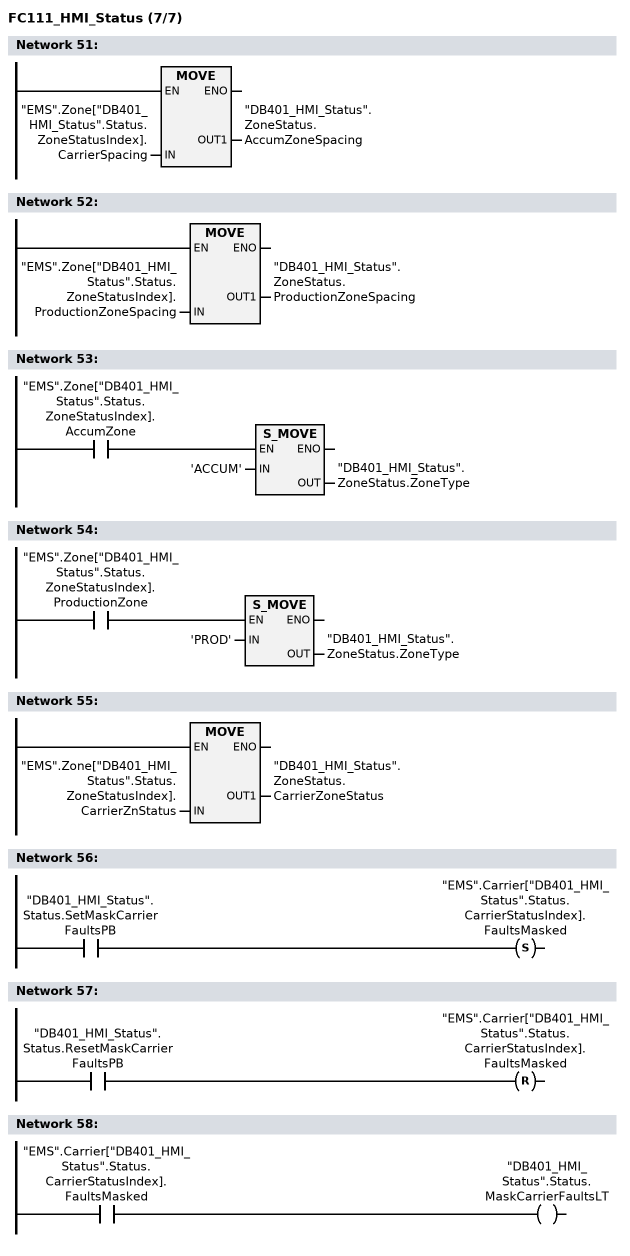
   RUNG wire#powerrail
      Move(in := "EMS".Zone["DB401_HMI_Status".Status.ZoneStatusIndex].CarrierSpacing, out1 => "DB401_HMI_Status".ZoneStatus.AccumZoneSpacing)
   END_RUNG
   // the same network as SCL:
   "DB401_HMI_Status".ZoneStatus.AccumZoneSpacing := "EMS".Zone["DB401_HMI_Status".Status.ZoneStatusIndex].CarrierSpacing;
END_REGION

REGION Network 52
   RUNG wire#powerrail
      Move(in := "EMS".Zone["DB401_HMI_Status".Status.ZoneStatusIndex].ProductionZoneSpacing, out1 => "DB401_HMI_Status".ZoneStatus.ProductionZoneSpacing)
   END_RUNG
   // the same network as SCL:
   "DB401_HMI_Status".ZoneStatus.ProductionZoneSpacing := "EMS".Zone["DB401_HMI_Status".Status.ZoneStatusIndex].ProductionZoneSpacing;
END_REGION

REGION Network 53
   RUNG wire#powerrail
      Contact( "EMS".Zone["DB401_HMI_Status".Status.ZoneStatusIndex].AccumZone )
      S_Move(in := 'ACCUM', out => "DB401_HMI_Status".ZoneStatus.ZoneType)
   END_RUNG
   // the same network as SCL:
   IF "EMS".Zone["DB401_HMI_Status".Status.ZoneStatusIndex].AccumZone THEN
       "DB401_HMI_Status".ZoneStatus.ZoneType := 'ACCUM';
   END_IF;
END_REGION

REGION Network 54
   RUNG wire#powerrail
      Contact( "EMS".Zone["DB401_HMI_Status".Status.ZoneStatusIndex].ProductionZone )
      S_Move(in := 'PROD', out => "DB401_HMI_Status".ZoneStatus.ZoneType)
   END_RUNG
   // the same network as SCL:
   IF "EMS".Zone["DB401_HMI_Status".Status.ZoneStatusIndex].ProductionZone THEN
       "DB401_HMI_Status".ZoneStatus.ZoneType := 'PROD';
   END_IF;
END_REGION

REGION Network 55
   RUNG wire#powerrail
      Move(in := "EMS".Zone["DB401_HMI_Status".Status.ZoneStatusIndex].CarrierZnStatus, out1 => "DB401_HMI_Status".ZoneStatus.CarrierZoneStatus)
   END_RUNG
   // the same network as SCL:
   "DB401_HMI_Status".ZoneStatus.CarrierZoneStatus := "EMS".Zone["DB401_HMI_Status".Status.ZoneStatusIndex].CarrierZnStatus;
END_REGION

REGION Network 56
   RUNG wire#powerrail
      Contact( "DB401_HMI_Status".Status.SetMaskCarrierFaultsPB )
      S_Coil( "EMS".Carrier["DB401_HMI_Status".Status.CarrierStatusIndex].FaultsMasked )
   END_RUNG
   // the same network as SCL:
   IF "DB401_HMI_Status".Status.SetMaskCarrierFaultsPB THEN
       "EMS".Carrier["DB401_HMI_Status".Status.CarrierStatusIndex].FaultsMasked := TRUE;
   END_IF;
END_REGION

REGION Network 57
   RUNG wire#powerrail
      Contact( "DB401_HMI_Status".Status.ResetMaskCarrierFaultsPB )
      R_Coil( "EMS".Carrier["DB401_HMI_Status".Status.CarrierStatusIndex].FaultsMasked )
   END_RUNG
   // the same network as SCL:
   IF "DB401_HMI_Status".Status.ResetMaskCarrierFaultsPB THEN
       "EMS".Carrier["DB401_HMI_Status".Status.CarrierStatusIndex].FaultsMasked := FALSE;
   END_IF;
END_REGION

REGION Network 58
   RUNG wire#powerrail
      Contact( "EMS".Carrier["DB401_HMI_Status".Status.CarrierStatusIndex].FaultsMasked )
      Coil( "DB401_HMI_Status".Status.MaskCarrierFaultsLT )
   END_RUNG
   // the same network as SCL:
   "DB401_HMI_Status".Status.MaskCarrierFaultsLT := "EMS".Carrier["DB401_HMI_Status".Status.CarrierStatusIndex].FaultsMasked;
END_REGION
END_FUNCTION

FUNCTION "FC201_SDC_To_Carrier_Map_IO [C01-C10]" : Void   // FC201, LAD
{ S7_Optimized_Access := 'TRUE' }
VERSION : 0.1
   VAR_TEMP
      templatch : Bool;
   END_VAR
BEGIN

REGION Network 1
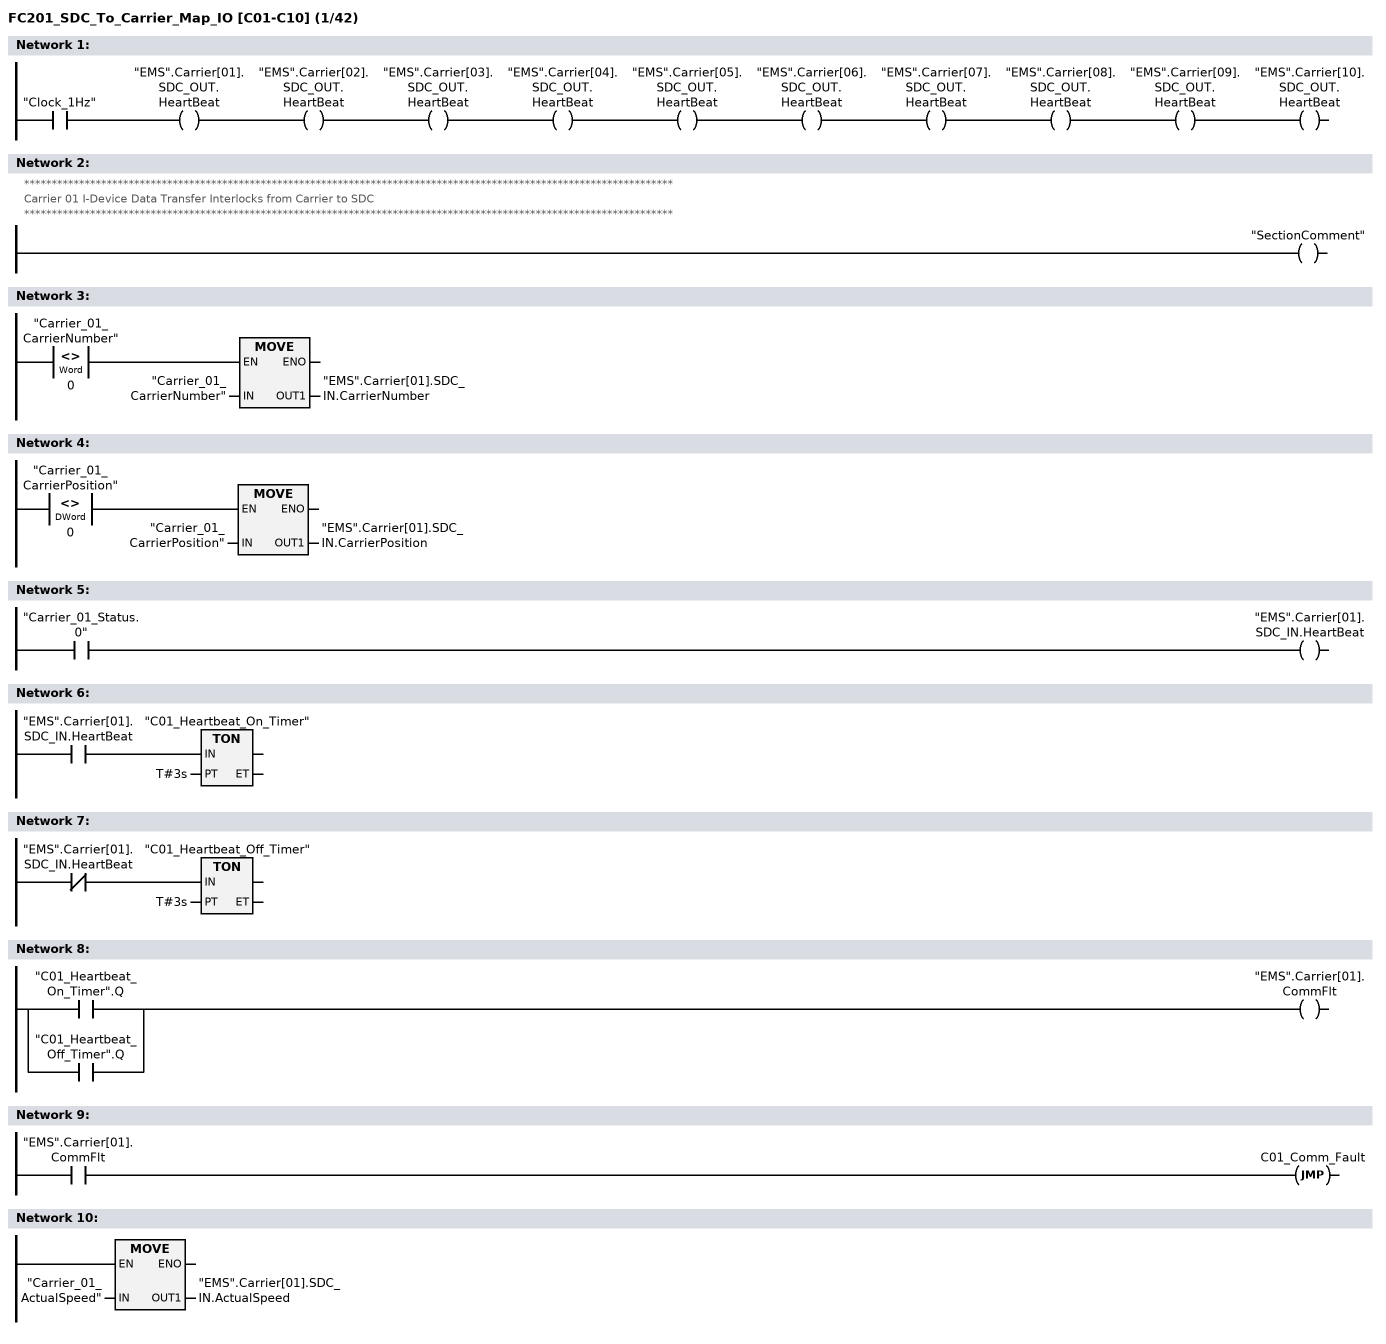
   RUNG wire#powerrail
      Contact( "Clock_1Hz" )
      Coil( "EMS".Carrier[01].SDC_OUT.HeartBeat )
      Coil( "EMS".Carrier[02].SDC_OUT.HeartBeat )
      Coil( "EMS".Carrier[03].SDC_OUT.HeartBeat )
      Coil( "EMS".Carrier[04].SDC_OUT.HeartBeat )
      Coil( "EMS".Carrier[05].SDC_OUT.HeartBeat )
      Coil( "EMS".Carrier[06].SDC_OUT.HeartBeat )
      Coil( "EMS".Carrier[07].SDC_OUT.HeartBeat )
      Coil( "EMS".Carrier[08].SDC_OUT.HeartBeat )
      Coil( "EMS".Carrier[09].SDC_OUT.HeartBeat )
      Coil( "EMS".Carrier[10].SDC_OUT.HeartBeat )
   END_RUNG
   // the same network as SCL:
   "EMS".Carrier[01].SDC_OUT.HeartBeat := "Clock_1Hz";
   "EMS".Carrier[02].SDC_OUT.HeartBeat := "Clock_1Hz";
   "EMS".Carrier[03].SDC_OUT.HeartBeat := "Clock_1Hz";
   "EMS".Carrier[04].SDC_OUT.HeartBeat := "Clock_1Hz";
   "EMS".Carrier[05].SDC_OUT.HeartBeat := "Clock_1Hz";
   "EMS".Carrier[06].SDC_OUT.HeartBeat := "Clock_1Hz";
   "EMS".Carrier[07].SDC_OUT.HeartBeat := "Clock_1Hz";
   "EMS".Carrier[08].SDC_OUT.HeartBeat := "Clock_1Hz";
   "EMS".Carrier[09].SDC_OUT.HeartBeat := "Clock_1Hz";
   "EMS".Carrier[10].SDC_OUT.HeartBeat := "Clock_1Hz";
END_REGION

REGION Network 2
   // **********************************************************************************************************************
   // 
   // Carrier 01 I-Device Data Transfer Interlocks from Carrier to SDC
   // 
   // **********************************************************************************************************************
   RUNG wire#powerrail
      Coil( "SectionComment" )
   END_RUNG
   // the same network as SCL:
   "SectionComment" := TRUE;
END_REGION

REGION Network 3
   RUNG wire#powerrail
      { S7_Templates := "SrcType := Word" } NE_Contact(in1 := "Carrier_01_CarrierNumber", in2 := 0)
      Move(in := "Carrier_01_CarrierNumber", out1 => "EMS".Carrier[01].SDC_IN.CarrierNumber)
   END_RUNG
   // the same network as SCL:
   IF "Carrier_01_CarrierNumber" <> 0 THEN
       "EMS".Carrier[01].SDC_IN.CarrierNumber := "Carrier_01_CarrierNumber";
   END_IF;
END_REGION

REGION Network 4
   RUNG wire#powerrail
      { S7_Templates := "SrcType := DWord" } NE_Contact(in1 := "Carrier_01_CarrierPosition", in2 := 0)
      Move(in := "Carrier_01_CarrierPosition", out1 => "EMS".Carrier[01].SDC_IN.CarrierPosition)
   END_RUNG
   // the same network as SCL:
   IF "Carrier_01_CarrierPosition" <> 0 THEN
       "EMS".Carrier[01].SDC_IN.CarrierPosition := "Carrier_01_CarrierPosition";
   END_IF;
END_REGION

REGION Network 5
   RUNG wire#powerrail
      Contact( "Carrier_01_Status.0" )
      Coil( "EMS".Carrier[01].SDC_IN.HeartBeat )
   END_RUNG
   // the same network as SCL:
   "EMS".Carrier[01].SDC_IN.HeartBeat := "Carrier_01_Status.0";
END_REGION

REGION Network 6
   "C01_Heartbeat_On_Timer".TON(IN := "EMS".Carrier[01].SDC_IN.HeartBeat, PT := T#3s);
END_REGION

REGION Network 7
   "C01_Heartbeat_Off_Timer".TON(IN := NOT "EMS".Carrier[01].SDC_IN.HeartBeat, PT := T#3s);
END_REGION

REGION Network 8
   RUNG wire#powerrail
      Contact( "C01_Heartbeat_On_Timer".Q )
      wire#w1
      Coil( "EMS".Carrier[01].CommFlt )
   END_RUNG
   RUNG wire#powerrail
      Contact( "C01_Heartbeat_Off_Timer".Q )
   END_RUNG wire#w1
   // the same network as SCL:
   "EMS".Carrier[01].CommFlt := "C01_Heartbeat_On_Timer".Q OR "C01_Heartbeat_Off_Timer".Q;
END_REGION

REGION Network 9
   RUNG wire#powerrail
      Contact( "EMS".Carrier[01].CommFlt )
      JumpCoil( C01_Comm_Fault )
   END_RUNG
   // the same network as SCL:
   IF "EMS".Carrier[01].CommFlt THEN GOTO C01_Comm_Fault; END_IF;
END_REGION

REGION Network 10
   RUNG wire#powerrail
      Move(in := "Carrier_01_ActualSpeed", out1 => "EMS".Carrier[01].SDC_IN.ActualSpeed)
   END_RUNG
   // the same network as SCL:
   "EMS".Carrier[01].SDC_IN.ActualSpeed := "Carrier_01_ActualSpeed";
END_REGION

REGION Network 11
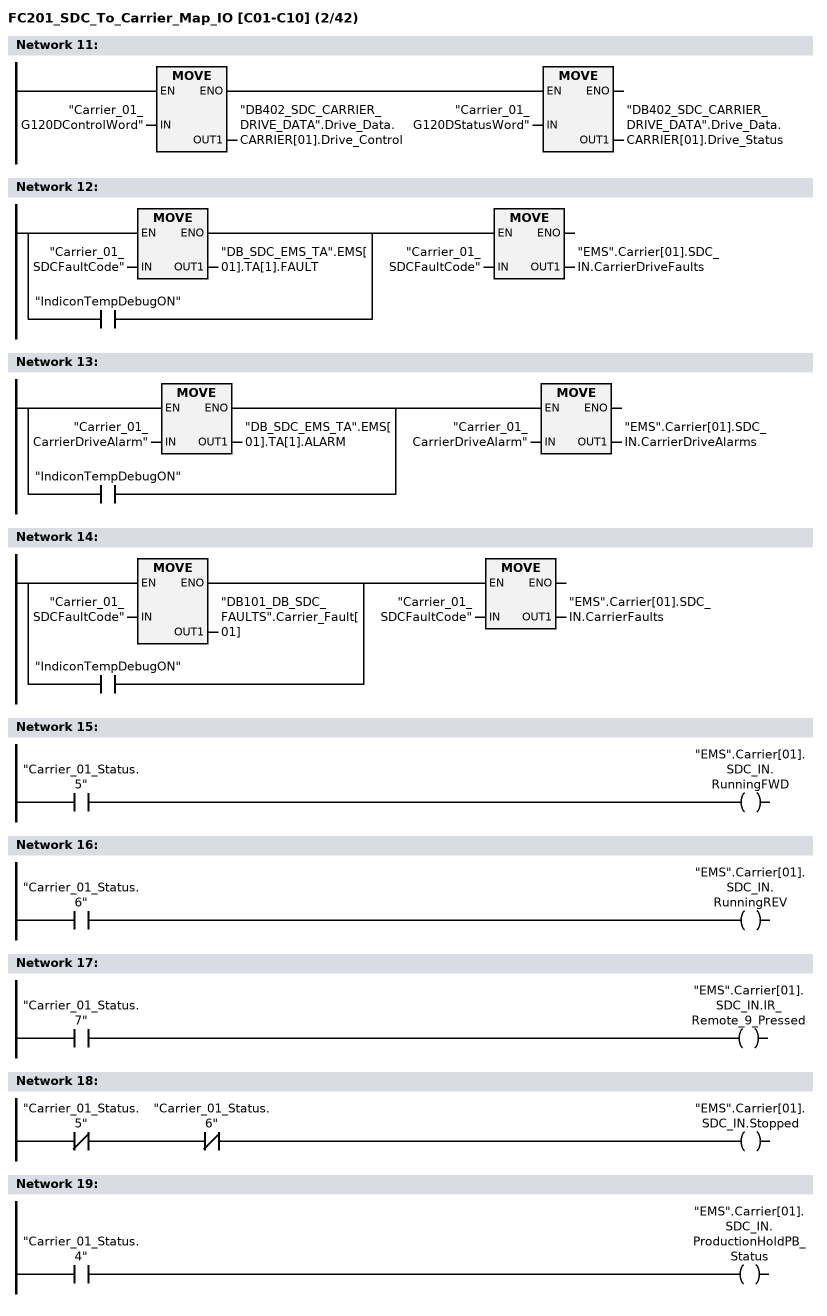
   RUNG wire#powerrail
      Move(in := "Carrier_01_G120DControlWord", out1 => "DB402_SDC_CARRIER_DRIVE_DATA".Drive_Data.CARRIER[01].Drive_Control)
      Move(in := "Carrier_01_G120DStatusWord", out1 => "DB402_SDC_CARRIER_DRIVE_DATA".Drive_Data.CARRIER[01].Drive_Status)
   END_RUNG
   // the same network as SCL:
   "DB402_SDC_CARRIER_DRIVE_DATA".Drive_Data.CARRIER[01].Drive_Control := "Carrier_01_G120DControlWord";
   "DB402_SDC_CARRIER_DRIVE_DATA".Drive_Data.CARRIER[01].Drive_Status := "Carrier_01_G120DStatusWord";
END_REGION

REGION Network 12
   RUNG wire#powerrail
      Move(in := "Carrier_01_SDCFaultCode", out1 => "DB_SDC_EMS_TA".EMS[01].TA[1].FAULT)
      wire#w1
      Move(in := "Carrier_01_SDCFaultCode", out1 => "EMS".Carrier[01].SDC_IN.CarrierDriveFaults)
   END_RUNG
   RUNG wire#powerrail
      Contact( "IndiconTempDebugON" )
   END_RUNG wire#w1
   // the same network as SCL:
   "DB_SDC_EMS_TA".EMS[01].TA[1].FAULT := "Carrier_01_SDCFaultCode";
   IF TRUE OR "IndiconTempDebugON" THEN
       "EMS".Carrier[01].SDC_IN.CarrierDriveFaults := "Carrier_01_SDCFaultCode";
   END_IF;
END_REGION

REGION Network 13
   RUNG wire#powerrail
      Move(in := "Carrier_01_CarrierDriveAlarm", out1 => "DB_SDC_EMS_TA".EMS[01].TA[1].ALARM)
      wire#w1
      Move(in := "Carrier_01_CarrierDriveAlarm", out1 => "EMS".Carrier[01].SDC_IN.CarrierDriveAlarms)
   END_RUNG
   RUNG wire#powerrail
      Contact( "IndiconTempDebugON" )
   END_RUNG wire#w1
   // the same network as SCL:
   "DB_SDC_EMS_TA".EMS[01].TA[1].ALARM := "Carrier_01_CarrierDriveAlarm";
   IF TRUE OR "IndiconTempDebugON" THEN
       "EMS".Carrier[01].SDC_IN.CarrierDriveAlarms := "Carrier_01_CarrierDriveAlarm";
   END_IF;
END_REGION

REGION Network 14
   RUNG wire#powerrail
      Move(in := "Carrier_01_SDCFaultCode", out1 => "DB101_DB_SDC_FAULTS".Carrier_Fault[01])
      wire#w1
      Move(in := "Carrier_01_SDCFaultCode", out1 => "EMS".Carrier[01].SDC_IN.CarrierFaults)
   END_RUNG
   RUNG wire#powerrail
      Contact( "IndiconTempDebugON" )
   END_RUNG wire#w1
   // the same network as SCL:
   "DB101_DB_SDC_FAULTS".Carrier_Fault[01] := "Carrier_01_SDCFaultCode";
   IF TRUE OR "IndiconTempDebugON" THEN
       "EMS".Carrier[01].SDC_IN.CarrierFaults := "Carrier_01_SDCFaultCode";
   END_IF;
END_REGION

REGION Network 15
   RUNG wire#powerrail
      Contact( "Carrier_01_Status.5" )
      Coil( "EMS".Carrier[01].SDC_IN.RunningFWD )
   END_RUNG
   // the same network as SCL:
   "EMS".Carrier[01].SDC_IN.RunningFWD := "Carrier_01_Status.5";
END_REGION

REGION Network 16
   RUNG wire#powerrail
      Contact( "Carrier_01_Status.6" )
      Coil( "EMS".Carrier[01].SDC_IN.RunningREV )
   END_RUNG
   // the same network as SCL:
   "EMS".Carrier[01].SDC_IN.RunningREV := "Carrier_01_Status.6";
END_REGION

REGION Network 17
   RUNG wire#powerrail
      Contact( "Carrier_01_Status.7" )
      Coil( "EMS".Carrier[01].SDC_IN.IR_Remote_9_Pressed )
   END_RUNG
   // the same network as SCL:
   "EMS".Carrier[01].SDC_IN.IR_Remote_9_Pressed := "Carrier_01_Status.7";
END_REGION

REGION Network 18
   RUNG wire#powerrail
      I_Contact( "Carrier_01_Status.5" )
      I_Contact( "Carrier_01_Status.6" )
      Coil( "EMS".Carrier[01].SDC_IN.Stopped )
   END_RUNG
   // the same network as SCL:
   "EMS".Carrier[01].SDC_IN.Stopped := NOT "Carrier_01_Status.5" AND NOT "Carrier_01_Status.6";
END_REGION

REGION Network 19
   RUNG wire#powerrail
      Contact( "Carrier_01_Status.4" )
      Coil( "EMS".Carrier[01].SDC_IN.ProductionHoldPB_Status )
   END_RUNG
   // the same network as SCL:
   "EMS".Carrier[01].SDC_IN.ProductionHoldPB_Status := "Carrier_01_Status.4";
END_REGION

REGION Network 20
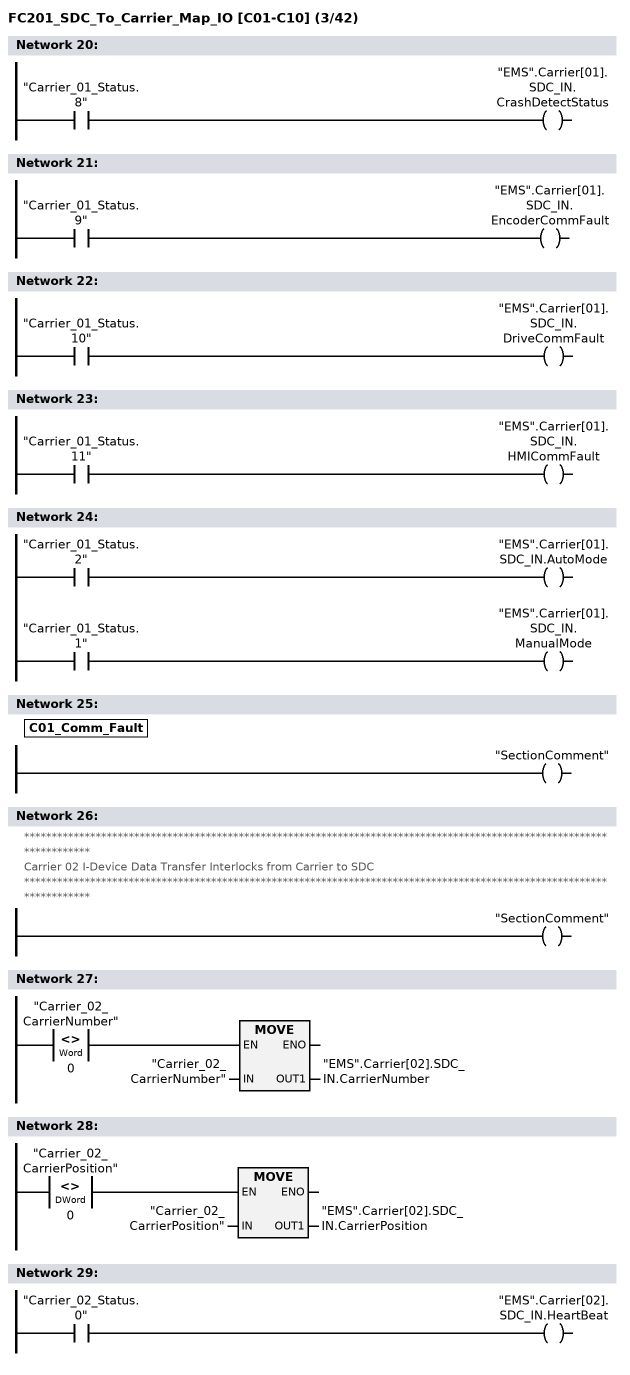
   RUNG wire#powerrail
      Contact( "Carrier_01_Status.8" )
      Coil( "EMS".Carrier[01].SDC_IN.CrashDetectStatus )
   END_RUNG
   // the same network as SCL:
   "EMS".Carrier[01].SDC_IN.CrashDetectStatus := "Carrier_01_Status.8";
END_REGION

REGION Network 21
   RUNG wire#powerrail
      Contact( "Carrier_01_Status.9" )
      Coil( "EMS".Carrier[01].SDC_IN.EncoderCommFault )
   END_RUNG
   // the same network as SCL:
   "EMS".Carrier[01].SDC_IN.EncoderCommFault := "Carrier_01_Status.9";
END_REGION

REGION Network 22
   RUNG wire#powerrail
      Contact( "Carrier_01_Status.10" )
      Coil( "EMS".Carrier[01].SDC_IN.DriveCommFault )
   END_RUNG
   // the same network as SCL:
   "EMS".Carrier[01].SDC_IN.DriveCommFault := "Carrier_01_Status.10";
END_REGION

REGION Network 23
   RUNG wire#powerrail
      Contact( "Carrier_01_Status.11" )
      Coil( "EMS".Carrier[01].SDC_IN.HMICommFault )
   END_RUNG
   // the same network as SCL:
   "EMS".Carrier[01].SDC_IN.HMICommFault := "Carrier_01_Status.11";
END_REGION

REGION Network 24
   RUNG wire#powerrail
      Contact( "Carrier_01_Status.2" )
      Coil( "EMS".Carrier[01].SDC_IN.AutoMode )
   END_RUNG
   RUNG wire#powerrail
      Contact( "Carrier_01_Status.1" )
      Coil( "EMS".Carrier[01].SDC_IN.ManualMode )
   END_RUNG
   // the same network as SCL:
   "EMS".Carrier[01].SDC_IN.AutoMode := "Carrier_01_Status.2";
   "EMS".Carrier[01].SDC_IN.ManualMode := "Carrier_01_Status.1";
END_REGION

REGION Network 25
   Label( C01_Comm_Fault )
   RUNG wire#powerrail
      Coil( "SectionComment" )
   END_RUNG
   // the same network as SCL:
   C01_Comm_Fault:
   "SectionComment" := TRUE;
END_REGION

REGION Network 26
   // **********************************************************************************************************************
   // 
   // Carrier 02 I-Device Data Transfer Interlocks from Carrier to SDC
   // 
   // **********************************************************************************************************************
   RUNG wire#powerrail
      Coil( "SectionComment" )
   END_RUNG
   // the same network as SCL:
   "SectionComment" := TRUE;
END_REGION

REGION Network 27
   RUNG wire#powerrail
      { S7_Templates := "SrcType := Word" } NE_Contact(in1 := "Carrier_02_CarrierNumber", in2 := 0)
      Move(in := "Carrier_02_CarrierNumber", out1 => "EMS".Carrier[02].SDC_IN.CarrierNumber)
   END_RUNG
   // the same network as SCL:
   IF "Carrier_02_CarrierNumber" <> 0 THEN
       "EMS".Carrier[02].SDC_IN.CarrierNumber := "Carrier_02_CarrierNumber";
   END_IF;
END_REGION

REGION Network 28
   RUNG wire#powerrail
      { S7_Templates := "SrcType := DWord" } NE_Contact(in1 := "Carrier_02_CarrierPosition", in2 := 0)
      Move(in := "Carrier_02_CarrierPosition", out1 => "EMS".Carrier[02].SDC_IN.CarrierPosition)
   END_RUNG
   // the same network as SCL:
   IF "Carrier_02_CarrierPosition" <> 0 THEN
       "EMS".Carrier[02].SDC_IN.CarrierPosition := "Carrier_02_CarrierPosition";
   END_IF;
END_REGION

REGION Network 29
   RUNG wire#powerrail
      Contact( "Carrier_02_Status.0" )
      Coil( "EMS".Carrier[02].SDC_IN.HeartBeat )
   END_RUNG
   // the same network as SCL:
   "EMS".Carrier[02].SDC_IN.HeartBeat := "Carrier_02_Status.0";
END_REGION

REGION Network 30
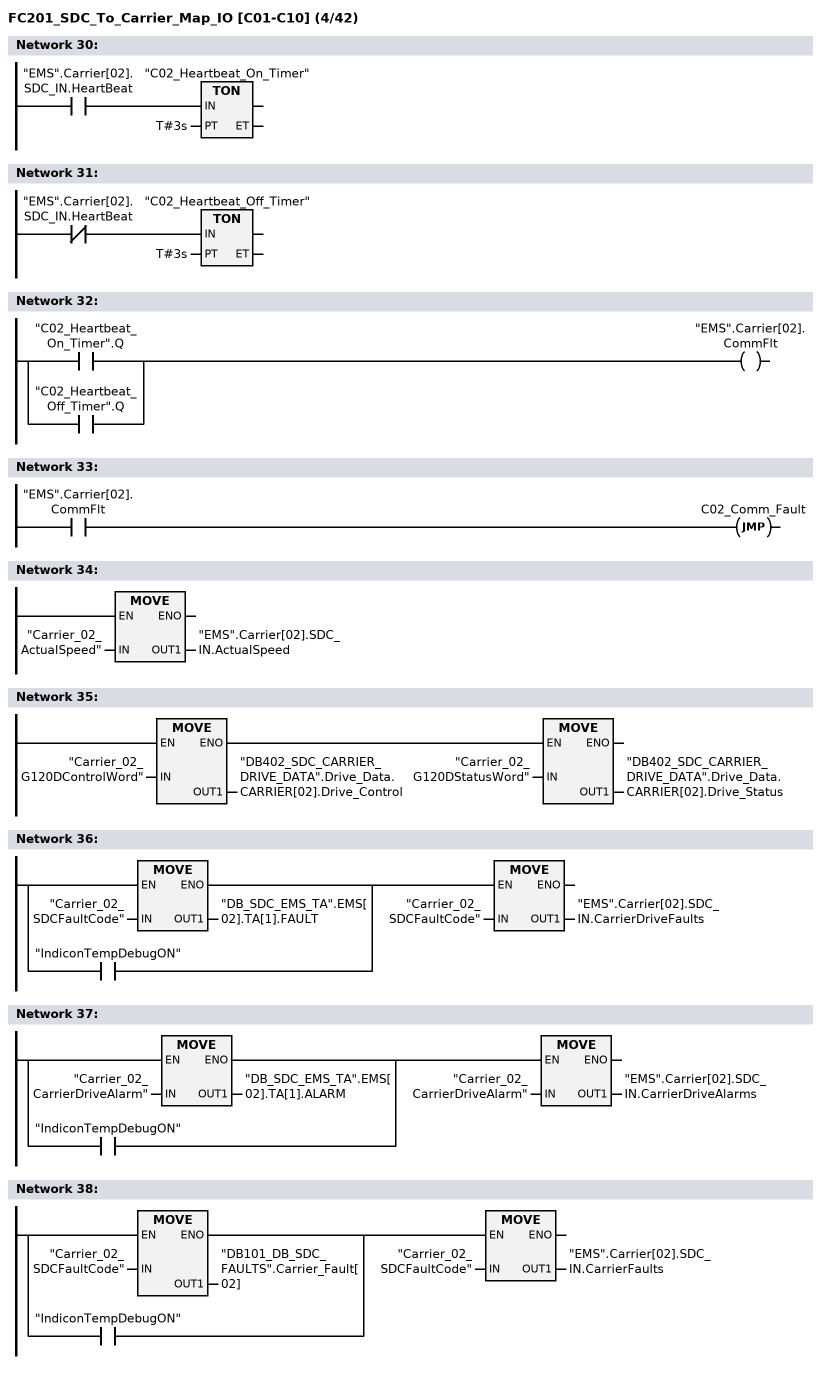
   "C02_Heartbeat_On_Timer".TON(IN := "EMS".Carrier[02].SDC_IN.HeartBeat, PT := T#3s);
END_REGION

REGION Network 31
   "C02_Heartbeat_Off_Timer".TON(IN := NOT "EMS".Carrier[02].SDC_IN.HeartBeat, PT := T#3s);
END_REGION

REGION Network 32
   RUNG wire#powerrail
      Contact( "C02_Heartbeat_On_Timer".Q )
      wire#w1
      Coil( "EMS".Carrier[02].CommFlt )
   END_RUNG
   RUNG wire#powerrail
      Contact( "C02_Heartbeat_Off_Timer".Q )
   END_RUNG wire#w1
   // the same network as SCL:
   "EMS".Carrier[02].CommFlt := "C02_Heartbeat_On_Timer".Q OR "C02_Heartbeat_Off_Timer".Q;
END_REGION

REGION Network 33
   RUNG wire#powerrail
      Contact( "EMS".Carrier[02].CommFlt )
      JumpCoil( C02_Comm_Fault )
   END_RUNG
   // the same network as SCL:
   IF "EMS".Carrier[02].CommFlt THEN GOTO C02_Comm_Fault; END_IF;
END_REGION

REGION Network 34
   RUNG wire#powerrail
      Move(in := "Carrier_02_ActualSpeed", out1 => "EMS".Carrier[02].SDC_IN.ActualSpeed)
   END_RUNG
   // the same network as SCL:
   "EMS".Carrier[02].SDC_IN.ActualSpeed := "Carrier_02_ActualSpeed";
END_REGION

REGION Network 35
   RUNG wire#powerrail
      Move(in := "Carrier_02_G120DControlWord", out1 => "DB402_SDC_CARRIER_DRIVE_DATA".Drive_Data.CARRIER[02].Drive_Control)
      Move(in := "Carrier_02_G120DStatusWord", out1 => "DB402_SDC_CARRIER_DRIVE_DATA".Drive_Data.CARRIER[02].Drive_Status)
   END_RUNG
   // the same network as SCL:
   "DB402_SDC_CARRIER_DRIVE_DATA".Drive_Data.CARRIER[02].Drive_Control := "Carrier_02_G120DControlWord";
   "DB402_SDC_CARRIER_DRIVE_DATA".Drive_Data.CARRIER[02].Drive_Status := "Carrier_02_G120DStatusWord";
END_REGION

REGION Network 36
   RUNG wire#powerrail
      Move(in := "Carrier_02_SDCFaultCode", out1 => "DB_SDC_EMS_TA".EMS[02].TA[1].FAULT)
      wire#w1
      Move(in := "Carrier_02_SDCFaultCode", out1 => "EMS".Carrier[02].SDC_IN.CarrierDriveFaults)
   END_RUNG
   RUNG wire#powerrail
      Contact( "IndiconTempDebugON" )
   END_RUNG wire#w1
   // the same network as SCL:
   "DB_SDC_EMS_TA".EMS[02].TA[1].FAULT := "Carrier_02_SDCFaultCode";
   IF TRUE OR "IndiconTempDebugON" THEN
       "EMS".Carrier[02].SDC_IN.CarrierDriveFaults := "Carrier_02_SDCFaultCode";
   END_IF;
END_REGION

REGION Network 37
   RUNG wire#powerrail
      Move(in := "Carrier_02_CarrierDriveAlarm", out1 => "DB_SDC_EMS_TA".EMS[02].TA[1].ALARM)
      wire#w1
      Move(in := "Carrier_02_CarrierDriveAlarm", out1 => "EMS".Carrier[02].SDC_IN.CarrierDriveAlarms)
   END_RUNG
   RUNG wire#powerrail
      Contact( "IndiconTempDebugON" )
   END_RUNG wire#w1
   // the same network as SCL:
   "DB_SDC_EMS_TA".EMS[02].TA[1].ALARM := "Carrier_02_CarrierDriveAlarm";
   IF TRUE OR "IndiconTempDebugON" THEN
       "EMS".Carrier[02].SDC_IN.CarrierDriveAlarms := "Carrier_02_CarrierDriveAlarm";
   END_IF;
END_REGION

REGION Network 38
   RUNG wire#powerrail
      Move(in := "Carrier_02_SDCFaultCode", out1 => "DB101_DB_SDC_FAULTS".Carrier_Fault[02])
      wire#w1
      Move(in := "Carrier_02_SDCFaultCode", out1 => "EMS".Carrier[02].SDC_IN.CarrierFaults)
   END_RUNG
   RUNG wire#powerrail
      Contact( "IndiconTempDebugON" )
   END_RUNG wire#w1
   // the same network as SCL:
   "DB101_DB_SDC_FAULTS".Carrier_Fault[02] := "Carrier_02_SDCFaultCode";
   IF TRUE OR "IndiconTempDebugON" THEN
       "EMS".Carrier[02].SDC_IN.CarrierFaults := "Carrier_02_SDCFaultCode";
   END_IF;
END_REGION

REGION Network 39
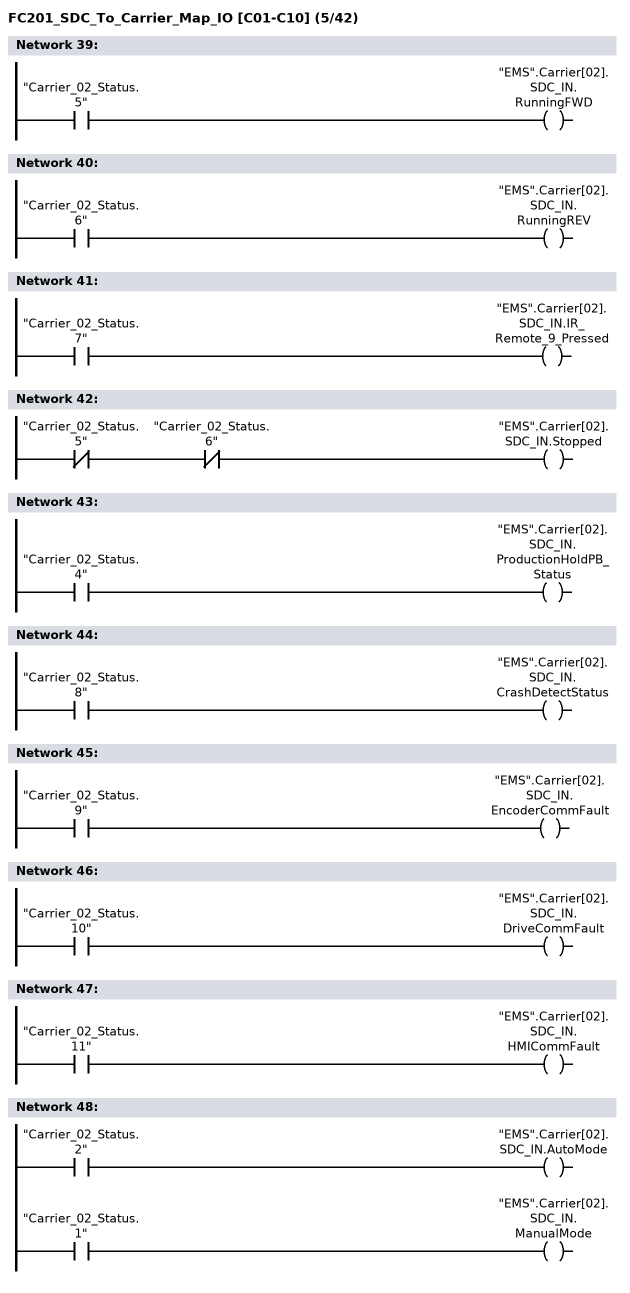
   RUNG wire#powerrail
      Contact( "Carrier_02_Status.5" )
      Coil( "EMS".Carrier[02].SDC_IN.RunningFWD )
   END_RUNG
   // the same network as SCL:
   "EMS".Carrier[02].SDC_IN.RunningFWD := "Carrier_02_Status.5";
END_REGION

REGION Network 40
   RUNG wire#powerrail
      Contact( "Carrier_02_Status.6" )
      Coil( "EMS".Carrier[02].SDC_IN.RunningREV )
   END_RUNG
   // the same network as SCL:
   "EMS".Carrier[02].SDC_IN.RunningREV := "Carrier_02_Status.6";
END_REGION

REGION Network 41
   RUNG wire#powerrail
      Contact( "Carrier_02_Status.7" )
      Coil( "EMS".Carrier[02].SDC_IN.IR_Remote_9_Pressed )
   END_RUNG
   // the same network as SCL:
   "EMS".Carrier[02].SDC_IN.IR_Remote_9_Pressed := "Carrier_02_Status.7";
END_REGION

REGION Network 42
   RUNG wire#powerrail
      I_Contact( "Carrier_02_Status.5" )
      I_Contact( "Carrier_02_Status.6" )
      Coil( "EMS".Carrier[02].SDC_IN.Stopped )
   END_RUNG
   // the same network as SCL:
   "EMS".Carrier[02].SDC_IN.Stopped := NOT "Carrier_02_Status.5" AND NOT "Carrier_02_Status.6";
END_REGION

REGION Network 43
   RUNG wire#powerrail
      Contact( "Carrier_02_Status.4" )
      Coil( "EMS".Carrier[02].SDC_IN.ProductionHoldPB_Status )
   END_RUNG
   // the same network as SCL:
   "EMS".Carrier[02].SDC_IN.ProductionHoldPB_Status := "Carrier_02_Status.4";
END_REGION

REGION Network 44
   RUNG wire#powerrail
      Contact( "Carrier_02_Status.8" )
      Coil( "EMS".Carrier[02].SDC_IN.CrashDetectStatus )
   END_RUNG
   // the same network as SCL:
   "EMS".Carrier[02].SDC_IN.CrashDetectStatus := "Carrier_02_Status.8";
END_REGION

REGION Network 45
   RUNG wire#powerrail
      Contact( "Carrier_02_Status.9" )
      Coil( "EMS".Carrier[02].SDC_IN.EncoderCommFault )
   END_RUNG
   // the same network as SCL:
   "EMS".Carrier[02].SDC_IN.EncoderCommFault := "Carrier_02_Status.9";
END_REGION

REGION Network 46
   RUNG wire#powerrail
      Contact( "Carrier_02_Status.10" )
      Coil( "EMS".Carrier[02].SDC_IN.DriveCommFault )
   END_RUNG
   // the same network as SCL:
   "EMS".Carrier[02].SDC_IN.DriveCommFault := "Carrier_02_Status.10";
END_REGION

REGION Network 47
   RUNG wire#powerrail
      Contact( "Carrier_02_Status.11" )
      Coil( "EMS".Carrier[02].SDC_IN.HMICommFault )
   END_RUNG
   // the same network as SCL:
   "EMS".Carrier[02].SDC_IN.HMICommFault := "Carrier_02_Status.11";
END_REGION

REGION Network 48
   RUNG wire#powerrail
      Contact( "Carrier_02_Status.2" )
      Coil( "EMS".Carrier[02].SDC_IN.AutoMode )
   END_RUNG
   RUNG wire#powerrail
      Contact( "Carrier_02_Status.1" )
      Coil( "EMS".Carrier[02].SDC_IN.ManualMode )
   END_RUNG
   // the same network as SCL:
   "EMS".Carrier[02].SDC_IN.AutoMode := "Carrier_02_Status.2";
   "EMS".Carrier[02].SDC_IN.ManualMode := "Carrier_02_Status.1";
END_REGION

REGION Network 49
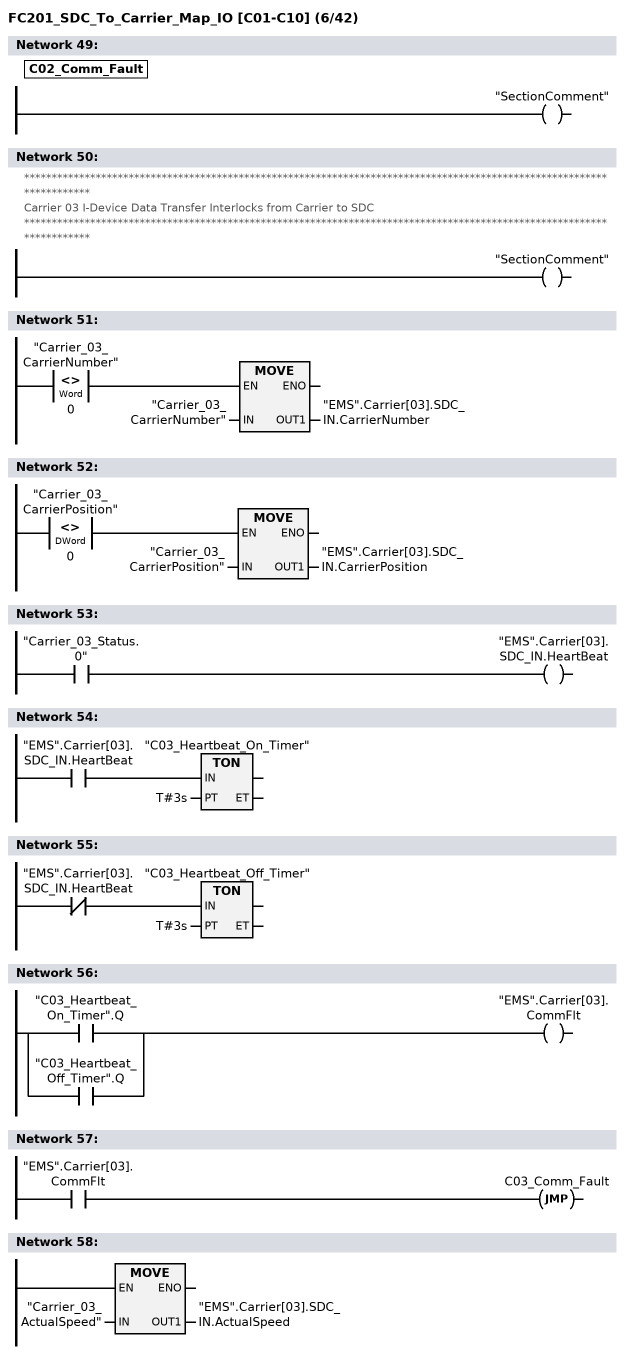
   Label( C02_Comm_Fault )
   RUNG wire#powerrail
      Coil( "SectionComment" )
   END_RUNG
   // the same network as SCL:
   C02_Comm_Fault:
   "SectionComment" := TRUE;
END_REGION

REGION Network 50
   // **********************************************************************************************************************
   // 
   // Carrier 03 I-Device Data Transfer Interlocks from Carrier to SDC
   // 
   // **********************************************************************************************************************
   RUNG wire#powerrail
      Coil( "SectionComment" )
   END_RUNG
   // the same network as SCL:
   "SectionComment" := TRUE;
END_REGION

REGION Network 51
   RUNG wire#powerrail
      { S7_Templates := "SrcType := Word" } NE_Contact(in1 := "Carrier_03_CarrierNumber", in2 := 0)
      Move(in := "Carrier_03_CarrierNumber", out1 => "EMS".Carrier[03].SDC_IN.CarrierNumber)
   END_RUNG
   // the same network as SCL:
   IF "Carrier_03_CarrierNumber" <> 0 THEN
       "EMS".Carrier[03].SDC_IN.CarrierNumber := "Carrier_03_CarrierNumber";
   END_IF;
END_REGION

REGION Network 52
   RUNG wire#powerrail
      { S7_Templates := "SrcType := DWord" } NE_Contact(in1 := "Carrier_03_CarrierPosition", in2 := 0)
      Move(in := "Carrier_03_CarrierPosition", out1 => "EMS".Carrier[03].SDC_IN.CarrierPosition)
   END_RUNG
   // the same network as SCL:
   IF "Carrier_03_CarrierPosition" <> 0 THEN
       "EMS".Carrier[03].SDC_IN.CarrierPosition := "Carrier_03_CarrierPosition";
   END_IF;
END_REGION

REGION Network 53
   RUNG wire#powerrail
      Contact( "Carrier_03_Status.0" )
      Coil( "EMS".Carrier[03].SDC_IN.HeartBeat )
   END_RUNG
   // the same network as SCL:
   "EMS".Carrier[03].SDC_IN.HeartBeat := "Carrier_03_Status.0";
END_REGION

REGION Network 54
   "C03_Heartbeat_On_Timer".TON(IN := "EMS".Carrier[03].SDC_IN.HeartBeat, PT := T#3s);
END_REGION

REGION Network 55
   "C03_Heartbeat_Off_Timer".TON(IN := NOT "EMS".Carrier[03].SDC_IN.HeartBeat, PT := T#3s);
END_REGION

REGION Network 56
   RUNG wire#powerrail
      Contact( "C03_Heartbeat_On_Timer".Q )
      wire#w1
      Coil( "EMS".Carrier[03].CommFlt )
   END_RUNG
   RUNG wire#powerrail
      Contact( "C03_Heartbeat_Off_Timer".Q )
   END_RUNG wire#w1
   // the same network as SCL:
   "EMS".Carrier[03].CommFlt := "C03_Heartbeat_On_Timer".Q OR "C03_Heartbeat_Off_Timer".Q;
END_REGION

REGION Network 57
   RUNG wire#powerrail
      Contact( "EMS".Carrier[03].CommFlt )
      JumpCoil( C03_Comm_Fault )
   END_RUNG
   // the same network as SCL:
   IF "EMS".Carrier[03].CommFlt THEN GOTO C03_Comm_Fault; END_IF;
END_REGION

REGION Network 58
   RUNG wire#powerrail
      Move(in := "Carrier_03_ActualSpeed", out1 => "EMS".Carrier[03].SDC_IN.ActualSpeed)
   END_RUNG
   // the same network as SCL:
   "EMS".Carrier[03].SDC_IN.ActualSpeed := "Carrier_03_ActualSpeed";
END_REGION

REGION Network 59
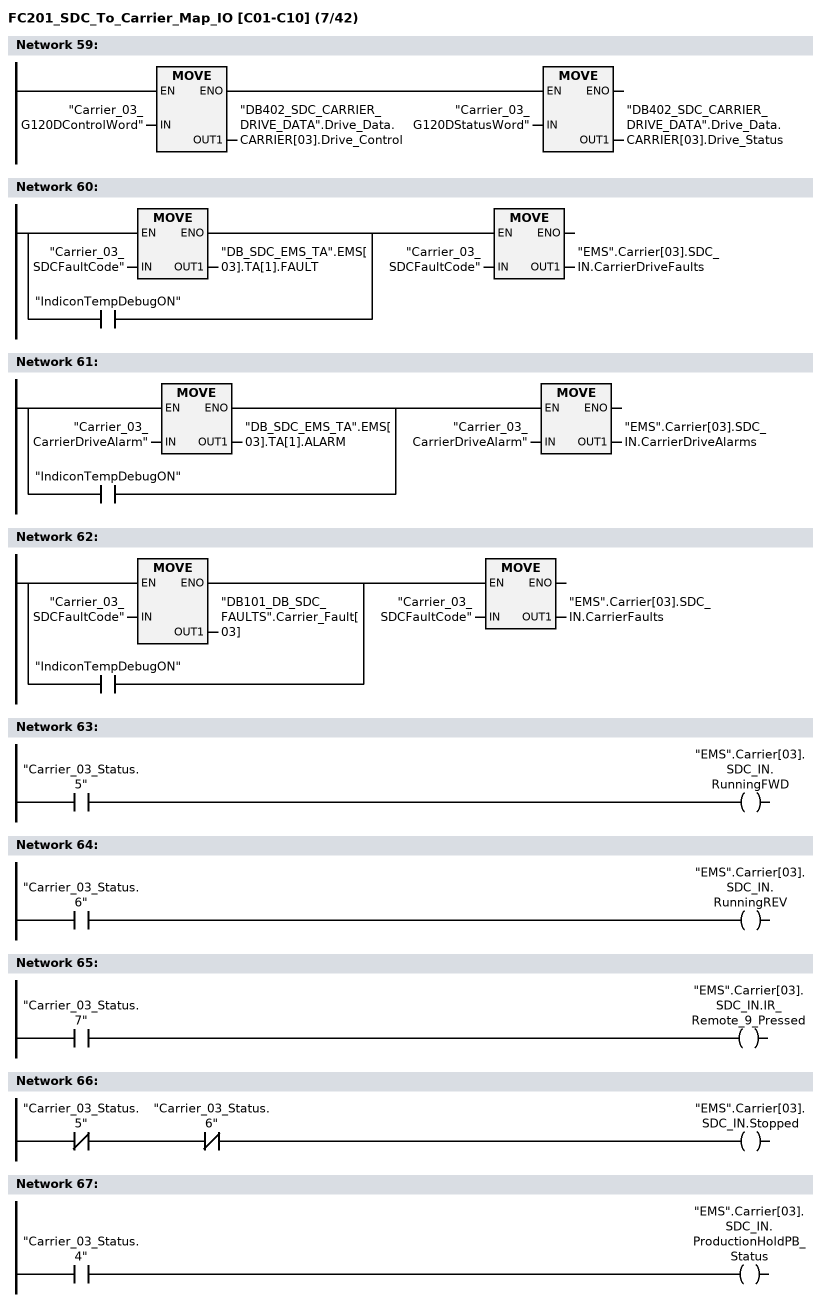
   RUNG wire#powerrail
      Move(in := "Carrier_03_G120DControlWord", out1 => "DB402_SDC_CARRIER_DRIVE_DATA".Drive_Data.CARRIER[03].Drive_Control)
      Move(in := "Carrier_03_G120DStatusWord", out1 => "DB402_SDC_CARRIER_DRIVE_DATA".Drive_Data.CARRIER[03].Drive_Status)
   END_RUNG
   // the same network as SCL:
   "DB402_SDC_CARRIER_DRIVE_DATA".Drive_Data.CARRIER[03].Drive_Control := "Carrier_03_G120DControlWord";
   "DB402_SDC_CARRIER_DRIVE_DATA".Drive_Data.CARRIER[03].Drive_Status := "Carrier_03_G120DStatusWord";
END_REGION

REGION Network 60
   RUNG wire#powerrail
      Move(in := "Carrier_03_SDCFaultCode", out1 => "DB_SDC_EMS_TA".EMS[03].TA[1].FAULT)
      wire#w1
      Move(in := "Carrier_03_SDCFaultCode", out1 => "EMS".Carrier[03].SDC_IN.CarrierDriveFaults)
   END_RUNG
   RUNG wire#powerrail
      Contact( "IndiconTempDebugON" )
   END_RUNG wire#w1
   // the same network as SCL:
   "DB_SDC_EMS_TA".EMS[03].TA[1].FAULT := "Carrier_03_SDCFaultCode";
   IF TRUE OR "IndiconTempDebugON" THEN
       "EMS".Carrier[03].SDC_IN.CarrierDriveFaults := "Carrier_03_SDCFaultCode";
   END_IF;
END_REGION
